(* Logix 5000 project; controller Digital_Interlock_PLC vendor 1 type 14 code 196 rev 37.11; software revision 37.00 *)

TASK MainTask (periodic, rate 10 ms, priority 5, watchdog 500 ms) : MainProgram

MODULES
   Local : vendor 1 type 14 code 196 (5069 0, rev 37.11)
      PF1 : vendor 1 type 14 code 107 (Ethernet 10.10.10.48, rev 37.1)
      ST1 : ETHERNET-MODULE (Ethernet 10.10.10.59, rev 1.1, Output RPI 10 ms)
           ST1:O.Data[0]   // To stacker heartbeat
           ST1:I.Data[1].0   // FeedInterruptStatus
      PR1 : ETHERNET-MODULE (Ethernet 10.10.10.6, rev 1.1, Output RPI 10 ms)
END_MODULES

TYPE STR_MajorFault :
STRUCT
   LEN : DINT;
   DATA : SINT[300];
END_STRUCT
END_TYPE

TYPE UDT_CommandEnum :
STRUCT
   cmd_none : DINT;
   cmd_start : DINT;
   cmd_stop : DINT;
   cmd_reset : DINT;
   cmd_interrupt : DINT;
   cmd_reconfigure : DINT;
END_STRUCT
END_TYPE

TYPE UDT_Constraints :
STRUCT
   GlobalSpeedMax : REAL;
   GlobalSpeedMin : REAL;
   KpiStabilityWindow_s : DINT;
END_STRUCT
END_TYPE

TYPE UDT_DeviceCmd :
STRUCT
   Mode : DINT;
   SpeedCmd : REAL;
   BufferTarget : DINT;
   Enable : BOOL;
END_STRUCT
END_TYPE

TYPE UDT_DeviceHealth :
STRUCT
   HeartbeatPrevious : BOOL;
   HeartbeartTimeout : BOOL;
   CommOK : BOOL;
   Enabled : BOOL;
   HeartbeatIn : BOOL;
   FaultInfo : DINT;
   EntryStatus : INT;
   FaultCode : INT;
   HBTimer : TIMER;
   Name : STRING;
   DeviceConfigured : BOOL;
END_STRUCT
END_TYPE

TYPE UDT_DeviceLink :
STRUCT
   ConnOK : BOOL;
   Simulation : BOOL;
   RoundTrip_ms : DINT;
   Handshake : UDT_Handshake;
   Cmd : UDT_DeviceCmd;
   Sts : UDT_DeviceSts;
END_STRUCT
END_TYPE

TYPE UDT_DeviceSts :
STRUCT
   PermissivesOK : BOOL;
   Running : BOOL;
   Faulted : BOOL;
   SpeedFB : REAL;
   BufferLevel : DINT;
   AlarmCode : DINT;
END_STRUCT
END_TYPE

TYPE UDT_DeviceTarget :
STRUCT
   DeviceID : DINT;
   SpeedMin : REAL;
   SpeedMax : REAL;
   BufferMin : DINT;
   BufferMax : DINT;
   Priority : DINT;
END_STRUCT
END_TYPE

TYPE UDT_EIP_DieCutter_FromStacker :   // Die cutter From Stacker
STRUCT
   blnFast : BOOL;   // Speed up die cutter (Stacker -> Press)
   blnSlow : BOOL;   // Slow down die cutter (Stacker -> Press)
   blnRegisterAdjustRq : BOOL;   // Move DC register to desired value (Stacker -> Press)
   blnRegisterStopAdjustRq : BOOL;   // Stop moving DC register (Stacker -> Press)
   blnSidewaysAdjustRq : BOOL;   // Move DC sideways to desired value (Stacker -> Press)
   blnSidewaysStopAdjustRq : BOOL;   // Stop DC sideways move (Stacker -> Press)
   blnSpeedChangeRq : BOOL;   // Change speed to desired speed (Stacker -> Press)
   blnSpeedChangeStopRq : BOOL;   // Stop speed change if active (Stacker -> Press)
   uiDesiredSpeedKpm : INT;   // 0-500 KPM (Stacker -> Press)
   fltDesiredRegisterAdjust : REAL;   // mm (Stacker -> Press)
   fltDesiredSidewaysAdjust : REAL;   // mm (Stacker -> Press)
END_STRUCT
END_TYPE

TYPE UDT_EIP_DieCutter_ToStacker :   // Die cutter to stacker
STRUCT
   blnRegistrationActive : BOOL;   // Die cutter registration motion active (Press -> Stacker)
   blnSidewaysAcitve : BOOL;   // Die cutter sideways motion active (Press -> Stacker)
   blnSpeedChangeActive : BOOL;   // Die cutter speed change active (Press -> Stacker)
   uiActualSpeedKpm : INT;   // Press current line speed (0-500 KPM) (Press -> Stacker)
   fltActualRegisterPosition : REAL;   // mm (Press -> Stacker)
   fltActualSidewaysPosition : REAL;   // mm (Press -> Stacker)
END_STRUCT
END_TYPE

TYPE UDT_EIP_FromBreaker :
STRUCT
   FeedInterrupted : BOOL;
   FeedInterrupt : BOOL;
   CurrentSpeed : DINT;
   CurrentFill : DINT;
   SampleRate : DINT;
   Deadband : DINT;
   MaxRunSpeed : DINT;
   MaxCmdSpeed : DINT;
   MinCmdSpeed : DINT;
   FeedInterruptSetting : DINT;
   TargetFill : DINT;
   CmdSpeed : DINT;
   Proportional : REAL;
   Name : STRING;
END_STRUCT
END_TYPE

TYPE UDT_EIP_FromConveyor :
STRUCT
   FeedInterrupt : BOOL;
   FeedInterrupted : BOOL;
   CurrentSpeed : DINT;
   CurrentFill : DINT;
   SampleRate : DINT;
   Deadband : DINT;
   MaxRunSpeed : DINT;
   MaxCmdSpeed : DINT;
   MinCmdSpeed : DINT;
   FeedInterruptSetting : DINT;
   TargetFill : DINT;
   CmdSpeed : DINT;
   Proportional : REAL;
   Name : STRING;
END_STRUCT
END_TYPE

TYPE UDT_EIP_FromPalletizer :
STRUCT
   FeedInterrupted : BOOL;
   FeedInterrupt : BOOL;
   CurrentSpeed : DINT;
   CurrentFill : DINT;
   SampleRate : DINT;
   Deadband : DINT;
   MaxRunSpeed : DINT;
   MaxCmdSpeed : DINT;
   MinCmdSpeed : DINT;
   FeedInterruptSetting : DINT;
   TargetFill : DINT;
   CmdSpeed : DINT;
   Proportional : REAL;
   Name : STRING;
END_STRUCT
END_TYPE

TYPE UDT_EIP_FromPrefeeder :
STRUCT
   AuxTamperAirRight : BOOL;   // (interlocks) (Pre-Feeder -> Press)
   AuxTamperAirLeft : BOOL;   // (interlocks) (Pre-Feeder -> Press)
   BackstopInhibit : BOOL;   // (Pre-Feeder -> Press)
   CallForStack : BOOL;   // Prefeeder calling for stack to be delivered (Prefeeder -> Floor Conv)
   ExtendoUpDown : BOOL;   // (interlocks) (Pre-Feeder -> Press)
   EstopFeedbackChannel1 : BOOL;   // (interlocks) (Pre-Feeder -> Press)
   EstopFeedbackChannel2 : BOOL;   // (interlocks) (Pre-Feeder -> Press)
   FeedBoardOk : BOOL;   // (interlocks) (Pre-Feeder -> Press)
   HeartbeatEcho : BOOL;
   MachineOpenCloseDisable : BOOL;   // (interlocks) (Pre-Feeder -> Press)
   OpenMachineOk : BOOL;   // (interlocks) (Pre-Feeder -> Press)
   ReadyForSetup : BOOL;   // (interlocks) (Pre-Feeder -> Press)
   ReadyToRaise : BOOL;   // (interlocks) (Pre-Feeder -> Press)
   RunEmpty : BOOL;   // (interlocks) (Pre-Feeder -> Press)
   RunForward : BOOL;   // Prefeeder telling conveyor to run forward (Prefeeder -> Floor Conv)
   RunReverse : BOOL;   // Prefeeder telling conveyor to run reverse (Prefeeder -> Floor Conv)
   TamperInterrupt : BOOL;   // (interlocks) (Pre-Feeder -> Press)
   CurrentSpeed : INT;   // Current speed of prefeeder (0-500KPM) (Pre-Feeder -> Press)
   PatternMaxSpeed : INT;   // Max speed allowed by stack pattern (0-500KPM) (Pre-Feeder -> Press)
END_STRUCT
END_TYPE

TYPE UDT_EIP_FromPress :
STRUCT
   ControlPowerInhibit : BOOL;   // Inhibit stacker from starting
   EstopOkChannel1 : BOOL;   // Press Estop is OK Ch1
   EstopOkChannel2 : BOOL;   // Press Estop is OK Ch2
   FeedEye : BOOL;   // Feed eye blocked (Press -> Stacker)
   GrinderCoverClosed : BOOL;   // OK to roll in
   LineSpeedSignal : DINT;   // Line speed of press (0-10V)
   LineEncoder : DINT;   // Enoder representing desired position of die cut cylinder rolls over every revolution (Press -> Stacker)
END_STRUCT
END_TYPE

TYPE UDT_EIP_FromStacker :
STRUCT
   ControlPower : BOOL;   // Stacker control power is on (interlocks)
   EstopOkChannel1 : BOOL;   // Stacker Estop to press ch1 (interlocks) (Stacker -> Press)
   EstopOkChannel2 : BOOL;   // Stacker Estop to press ch2 (interlocks) (Stacker -> Press)
   CompensatorControls : BOOL;   // Die Cut and Flexo Reg controls (interlocks)
   FeedInterruptStatus : BOOL;   // Interrupt request from stacker (status) (Stacker -> Press)
   FeedInterrupt : BOOL;   // Interrupt request from stacker (flow control) (Stacker -> Press)
   FeedRestart : BOOL;   // Restart feed (interlocks) (Stacker -> Press)
   HeartbeatEcho : BOOL;
   StackerRolledInChannel1 : BOOL;   // Stacker Rolled In to press Ok 2 Run Ch1 (interlocks) (Stacker -> Press)
   StackerRolledInChannel2 : BOOL;   // Stacker Rolled In to press Ok 2 Run Ch2 (interlocks) (Stacker -> Press)
   RunPermissive : BOOL;   // OK for press to run (interlocks) (Stacker -> Press)
   RolledOutStatus : BOOL;   // Die cutter rolled out (status) (Stacker -> Press)
   Spare1 : DINT;
   Spare2 : DINT;
   CurrentSpeed : INT;   // Current stacker line speed (0-500 KPM) (flow control) (Stacker -> Press)
   FillPercentage : INT;   // Percentage of Accumulation Consumed (for calculating Upstream Machine Speed) (flow control) (Stacker -> Press)
   PatternMaxSpeed : INT;   // Maximum speed allowed by stacker pattern (0-500 KPM) (flow control) (Stacker -> Press)
   Heartbeat : UINT;   // Heartbeat Reflection from Stacker (interlocks) (Stacker -> Press)
   DieCutter : UDT_EIP_DieCutter_FromStacker;
   PrintStation : UDT_EIP_PrintStation_FromStacker[7];
END_STRUCT
END_TYPE

TYPE UDT_EIP_FromStrapper :
STRUCT
   FeedInterrupt : BOOL;
   FeedInterrupted : BOOL;
   CurrentSpeed : DINT;
   CurrentFill : DINT;
   SampleRate : DINT;
   Deadband : DINT;
   MaxRunSpeed : DINT;
   MaxCmdSpeed : DINT;
   MinCmdSpeed : DINT;
   FeedInterruptSetting : DINT;
   TargetFill : DINT;
   CmdSpeed : DINT;
   Proportional : REAL;
   Name : STRING;
END_STRUCT
END_TYPE

TYPE UDT_EIP_FromTwinBoxSlitter :
STRUCT
   FeedInterrupt : BOOL;
   FeedInterrupted : BOOL;
   CurrentSpeed : DINT;
   CurrentFill : DINT;
   SampleRate : DINT;
   Deadband : DINT;
   MaxRunSpeed : DINT;
   MaxCmdSpeed : DINT;
   MinCmdSpeed : DINT;
   FeedInterruptSetting : DINT;
   TargetFill : DINT;
   CmdSpeed : DINT;
   Proportional : REAL;
   Name : STRING;
END_STRUCT
END_TYPE

TYPE UDT_EIP_PrintStation_FromStacker :   // print station from stacker
STRUCT
   blnRegisterAdjustRq : BOOL;   // (Stacker -> Press)
   blnSidewaysAdjustRq : BOOL;   // (Stacker -> Press)
   blnRegisterStopAdjustRq : BOOL;   // (Stacker -> Press)
   blnSidewaysStopAdjustRq : BOOL;   // (Stacker -> Press)
   fltDesiredRegisterAdjust : REAL;   // mm (Stacker -> Press)
   fltDesiredSidewaysAdjust : REAL;   // mm (Stacker -> Press)
END_STRUCT
END_TYPE

TYPE UDT_EIP_PrintStation_ToStacker :   // print station to stacker
STRUCT
   blnRegistrationActive : BOOL;   // (Press -> Stacker)
   blnSideWaysActive : BOOL;   // (Press -> Stacker)
   fltActualRegisterPosition : REAL;   // mm (Press -> Stacker)
   fltActualSidewaysPosition : REAL;   // mm (Press -> Stacker)
END_STRUCT
END_TYPE

TYPE UDT_EIP_ToBreaker :
STRUCT
   FeedInterrupted : BOOL;
   FeedInterrupt : BOOL;
   CurrentSpeed : DINT;
   CurrentFill : DINT;
   SampleRate : DINT;
   Deadband : DINT;
   MaxRunSpeed : DINT;
   MaxCmdSpeed : DINT;
   MinCmdSpeed : DINT;
   FeedInterruptSetting : DINT;
   TargetFill : DINT;
   CmdSpeed : DINT;
   Proportional : REAL;
   Name : STRING;
END_STRUCT
END_TYPE

TYPE UDT_EIP_ToConveyor :
STRUCT
   FeedInterrupt : BOOL;
   FeedInterrupted : BOOL;
   CurrentSpeed : DINT;
   CurrentFill : DINT;
   SampleRate : DINT;
   Deadband : DINT;
   MaxRunSpeed : DINT;
   MaxCmdSpeed : DINT;
   MinCmdSpeed : DINT;
   FeedInterruptSetting : DINT;
   TargetFill : DINT;
   CmdSpeed : DINT;
   Proportional : REAL;
   Name : STRING;
END_STRUCT
END_TYPE

TYPE UDT_EIP_ToPalletizer :
STRUCT
   FeedInterrupted : BOOL;
   FeedInterrupt : BOOL;
   CurrentSpeed : DINT;
   CurrentFill : DINT;
   SampleRate : DINT;
   Deadband : DINT;
   MaxRunSpeed : DINT;
   MaxCmdSpeed : DINT;
   MinCmdSpeed : DINT;
   FeedInterruptSetting : DINT;
   TargetFill : DINT;
   CmdSpeed : DINT;
   Proportional : REAL;
   Name : STRING;
END_STRUCT
END_TYPE

TYPE UDT_EIP_ToPrefeeder :
STRUCT
   ClosedLocked : BOOL;   // (interlocks) (Press -> Pre-Feeder)
   ConvRunning : BOOL;   // (Floor Conv -> Prefeeder)
   ExtendoFollowBackstopUp : BOOL;   // (interlocks) (Press -> Pre-Feeder)
   ExtendoFollowBackstopDown : BOOL;   // (interlocks) (Press -> Pre-Feeder)
   LastStack : BOOL;   // Last stack running in (Floor Conv -> Prefeeder)
   LoadHopper : BOOL;   // (interlocks) (Press -> Pre-Feeder)
   MachineInFeedMode : BOOL;   // (interlocks) (Press -> Pre-Feeder)
   MachineRunning : BOOL;   // (interlocks) (Press -> Pre-Feeder)
   RequestsOpen : BOOL;   // (interlocks) (Press -> Pre-Feeder)
   StackReadyInFeed : BOOL;   // Stack is present at the end of the floor conveyor (Floor Conv -> Prefeeder)
   ShuttleCarAtPrefeeder : BOOL;   // (Floor Conv -> Prefeeder)
   Heartbeat : DINT;
   CommandedSpeed : INT;   // Commanded speed from the Press/LIC (0-500KPM) (flow control) (Press -> Pre-Feeder)
   BoardCaliper : REAL;   // Thickness of board (mm) (interlocks) (Press -> Pre-Feeder)
   FeedHopperHeight : REAL;   // (mm) (interlocks) (Press -> Pre-Feeder)
   HopperHeightSetpoint : REAL;   // (mm) (interlocks) (Press -> Pre-Feeder)
   HopperHeightMin : REAL;   // (mm) (interlocks) (Press -> Pre-Feeder)
   LinearSpeedSetpoint : REAL;   // Setting based on recipe (mm/s) (interlocks) (Press -> Pre-Feeder)
   LinearSpeedActual : REAL;   // Actual speed (mm/s) (interlocks) (Press -> Pre-Feeder)
END_STRUCT
END_TYPE

TYPE UDT_EIP_ToPress :
STRUCT
   AuxTamperAirRight : BOOL;   // (Pre-Feeder -> Press)
   AuxTamperAirLeft : BOOL;   // (Pre-Feeder -> Press)
   CallForStack : BOOL;   // Prefeeder -> Floor Conv
   FeedBoardOk : BOOL;   // (Pre-Feeder -> Press)
   MachineOpenCloseDisable : BOOL;   // (Pre-Feeder -> Press)
   OpenMachineOk : BOOL;   // (Pre-Feeder -> Press)
   ReadyForSetup : BOOL;   // (Pre-Feeder -> Press)
   ReadyToRaise : BOOL;   // (Pre-Feeder -> Press)
   RunEmpty : BOOL;
   RunForward : BOOL;   // (Pre-Feeder -> Press)
   RunReverse : BOOL;   // (Pre-Feeder -> Press)
   TamperInterrupt : BOOL;   // (Pre-Feeder -> Press)
   Empty : BOOL;   // (Pre-Feeder -> Press)
   BackstopInhibit : BOOL;   // (Prefeeder -> Press)
   Placeholder : BOOL;
   FeedInterrupt : BOOL;   // Interrupt request from stacker (flow control)
   FeedRestart : BOOL;   // Restart feed (interlocks)
   EstopFeedbackChannel1 : BOOL;   // (Prefeeder -> Press)
   EstopFeedbackChannel2 : BOOL;   // (Prefeeder -> Press)
   EstopOkChannel1 : BOOL;   // Stacker Estop to press ch1 (interlocks)
   EstopOkChannel2 : BOOL;   // Stacker Estop to press ch2 (interlocks)
   ExtendoUpDown : BOOL;   // (interlocks) (Pre-Feeder -> Press)
   StackerRolledInChannel1 : BOOL;   // Stacker Rolled In to press Ok 2 Run Ch1 (interlocks)
   StackerRolledInChannel2 : BOOL;   // Stacker Rolled In to press Ok 2 Run Ch2 (interlocks)
   ControlPower : BOOL;   // Stacker control power is on (interlocks)
   CompensatorControls : BOOL;   // Die Cut and Flexo Reg controls (interlocks)
   RunPermissive : BOOL;   // OK for press to run (interlocks)
   RolledOutStatus : BOOL;   // Die cutter rolled out (status)
   FeedInterruptStatus : BOOL;   // Interrupt request from stacker (status)
   Spare : BOOL;
   Heartbeat_Echo_Prefeeder : UINT;   // Heartbeat Reflection from Prefeeder (interlocks) (Prefeeder -> Press)
   Heartbeat_Echo_Stacker : UINT;   // Heartbeat Reflection from Stacker (interlocks) (Stacker -> Press)
   CurrentSpeed : UINT;   // Current stacker line speed (0-500 KPM) (flow control) (Pre-Feeder -> Press)
   PatternMaxSpeed : UINT;   // Maximum speed allowed by stacker pattern (0-500 KPM) (flow control) (Pre-Feeder -> Press)
   FillPercentage : UINT;   // Percentage of Accumulation Consumed (for calculating Upstream Machine Speed) (flow control)
   Spare1 : DINT;
   Spare2 : DINT;
   DieCutter : UDT_EIP_DieCutter_ToStacker;
   PrintStation : UDT_EIP_PrintStation_FromStacker[7];
END_STRUCT
END_TYPE

TYPE UDT_EIP_ToStacker :
STRUCT
   ControlPowerInhibit : BOOL;   // ADDED FOR EIP COMMS Inhibit stacker from starting
   DownstreamReady : BOOL;   // (LIC -> Stacker)
   EstopOkChannel1 : BOOL;   // Press Estop is OK Ch1 (interlocks) (Press -> Stacker)
   EstopOkChannel2 : BOOL;   // Press Estop is OK Ch2 (interlocks) (Press -> Stacker)
   FeedEye : BOOL;   // ADDED FOR EIP COMMS Feed eye blocked
   GrinderCoverClosed : BOOL;   // ADDED FOR EIP COMMS OK to roll in
   RollInPermissive : BOOL;   // Permission for stacker roll-in (Press -> Stacker)
   RunPermissive : BOOL;   // Rum permissive from press (interlocks) (Press -> Stacker)
   SheetCountPulseStatus : BOOL;   // Sheet count pulse (interlocks) (Press -> Stacker)
   VOSReset : BOOL;   // Reset VOS faults (if applicable) (interlocks) (Press -> Stacker)
   VOSStart : BOOL;   // Start VOS (if applicable) (interlocks) (Press -> Stacker)
   CommsStatus : DINT;   // (Interlock -> Stacker)
   Spare1 : DINT;
   Spare2 : DINT;
   LineEncoder : DINT;   // ADDED FOR EIP COMMS Enoder representing desired position of die cut cylinder rolls over every revolution
   LineSpeedSignal : DINT;   // ADDED FOR EIP COMMS Line speed of press (0-10V)
   CommandedSpeed : INT;   // Commanded press speed (0-500 KPM) (Press -> Stacker)
   PressCurrentSpeed : INT;   // Actual press speed (0-500 KPM) (Press -> Stacker)
   Heartbeat : UINT;   // Incrementing heartbeat for comm health (Press -> Stacker)
   DieCutter : UDT_EIP_DieCutter_ToStacker;
   PrintStation : UDT_EIP_PrintStation_ToStacker[7];
END_STRUCT
END_TYPE

TYPE UDT_EIP_ToStrapper :
STRUCT
   FeedInterrupt : BOOL;
   FeedInterrupted : BOOL;
   CurrentSpeed : DINT;
   CurrentFill : DINT;
   SampleRate : DINT;
   Deadband : DINT;
   MaxRunSpeed : DINT;
   MaxCmdSpeed : DINT;
   MinCmdSpeed : DINT;
   FeedInterruptSetting : DINT;
   TargetFill : DINT;
   CmdSpeed : DINT;
   Proportional : REAL;
   Name : STRING;
END_STRUCT
END_TYPE

TYPE UDT_EIP_ToTwinBoxSlitter :
STRUCT
   FeedInterrupt : BOOL;
   FeedInterrupted : BOOL;
   CurrentSpeed : DINT;
   CurrentFill : DINT;
   SampleRate : DINT;
   Deadband : DINT;
   MaxRunSpeed : DINT;
   MaxCmdSpeed : DINT;
   MinCmdSpeed : DINT;
   FeedInterruptSetting : DINT;
   TargetFill : DINT;
   CmdSpeed : DINT;
   Proportional : REAL;
   Name : STRING;
END_STRUCT
END_TYPE

TYPE UDT_FaultRecord :
STRUCT
   TimeLow : DINT;
   TimeHigh : DINT;
   Type : INT;
   Code : INT;
   Info : DINT[11];
END_STRUCT
END_TYPE

TYPE UDT_FromLIC :   // Data that is exchanged with LIC Client
STRUCT
   EnableLineOptimization : BOOL;
   Deadband : DINT;
   FeedInterruptSetting : DINT;
   MaxCommandSpeed : DINT;
   MinCommandSpeed : DINT;
   Proportional : DINT;
   SampleRate : DINT;
   TargetFillPercentage : DINT;
   MachineList : STRING;
   ToBR1 : UDT_EIP_ToBreaker;
   ToBR2 : UDT_EIP_ToBreaker;
   ToCN1 : UDT_EIP_ToConveyor;
   ToCN2 : UDT_EIP_ToConveyor;
   ToPL1 : UDT_EIP_ToPalletizer;
   ToPL2 : UDT_EIP_ToPalletizer;
   ToFE1 : UDT_EIP_ToPrefeeder;
   ToFE2 : UDT_EIP_ToPrefeeder;
   ToPR1 : UDT_EIP_ToPress;
   ToPR2 : UDT_EIP_ToPress;
   ToST1 : UDT_EIP_ToStacker;
   ToST2 : UDT_EIP_ToStacker;
   ToTB1 : UDT_EIP_ToTwinBoxSlitter;
   ToTB2 : UDT_EIP_ToTwinBoxSlitter;
   ToSR1 : UDT_EIP_ToStrapper;
   ToSR2 : UDT_EIP_ToStrapper;
END_STRUCT
END_TYPE

TYPE UDT_GenericStacker :
STRUCT
   cmd : DINT;
   status : DINT;
END_STRUCT
END_TYPE

TYPE UDT_Handshake :   // Device handshake and telemetry
STRUCT
   Req : BOOL;
   Ack : BOOL;
   Busy : BOOL;
   Done : BOOL;
   Fault : BOOL;
   TxnID : DINT;
   TxnIDEcho : DINT;
   Timeout_ms : DINT;
   Timer_ms : DINT;
END_STRUCT
END_TYPE

TYPE UDT_MachineType :
STRUCT
   ModuleExists : BOOL;   // (Handled by SetModuleInhibitMode) A bool that represents unihibited (0,False) or inhibited (1,True)
   FeedInterrupt : BOOL;   // (Output to each PLC) Boolean for activating feed interrupt
   FeedInterrupted : BOOL;   // Flag to verify feed interrupt execution
   ProportialGain : REAL;   // Proportial multiple to adjust aggressiveness of changes to speed commands, limited to [0.5 - 1.2]
   MachineType : STRING;   // (From HMI) List of configured machines, with format "FE1,PR1,SR1,ST1,PL1"
   CurrentSpeed : DINT;   // (From each PLC) Each machine will have a current speed value, obtained over EIP
   MinSpeed : DINT;   // (From each PLC) Minimum speed of the machine
   CommandSpeed : DINT;   // (Output of Line Flow Opt) Commanded speed adjustment from speed algorithm, occurs every *evaluation interval*
   IPSubnet : DINT;   // (**CHECK** if HMI will provide) The subnet that maps to the type of machine
   FeedInterruptSetting : DINT;   // (Input from HMI) Value from 0 to 100% , above which the press feed interrupt is triggered
   ReferenceSpeed : DINT;   // (Obtained from reference list, derived from machine list) Speed reference of downstream machine
   CurrFillPercentage : DINT;   // (From each PLC) Fill percentage of current machine
   TargFillPercentage : DINT;   // (From HMI per machine) The target fill percentage that is used to calculate commanded speeds
   Deadband : DINT;   // Value that represents the amount of percentage points from target fill percentage that the current fill percentage must be before calculating command speed
   MaxCmdSpeed : DINT;   // (From HMI) Value in KPM representing the upper limit of the commanded speed to be output to the upstream machine
   MinCmdSpeed : DINT;   // (From HMI) Value in KPM representing the lower limit of the commanded speed to be output to the upstream machine
END_STRUCT
END_TYPE

TYPE UDT_Optimize_Command :
STRUCT
   Enable : BOOL;
   Request : BOOL;
   Cancel : BOOL;
   Reset : BOOL;
END_STRUCT
END_TYPE

TYPE UDT_Optimize_Config :
STRUCT
   RecipeID : DINT;
   Mode : DINT;
   Targets : UDT_DeviceTarget[15];
   Constraints : UDT_Constraints;
END_STRUCT
END_TYPE

TYPE UDT_Optimize_Status :
STRUCT
   Active : BOOL;
   Busy : BOOL;
   Complete : BOOL;
   Fault : BOOL;
   Step : DINT;
   Substep : DINT;
   TimeInState_ms : DINT;
   LastErrorCode : DINT;
   LastErrorText : DINT;
   TxnID : DINT;
END_STRUCT
END_TYPE

TYPE UDT_StateContext :
STRUCT
   AbortReq : BOOL;
   Alarm : BOOL;
   Busy : BOOL;
   Complete : BOOL;
   InitDone : BOOL;
   StateChanged : BOOL;
   StartRisingEdge : BOOL;
   StopRisingEdge : BOOL;
   ResetRisingEdge : BOOL;
   PreviousStart : BOOL;
   PreviousStop : BOOL;
   PreviousReset : BOOL;
   InterruptRisingEdge : BOOL;
   PreviousInterrupt : BOOL;
   PreviousDone : BOOL;
   DoneRisingEdge : BOOL;
   Previous : DINT;
   Current : DINT;
   EntryStamp : DINT;   // ms since power-up
   TimeInState_ms : DINT;
   Command : DINT;   // from HMI/mailbox
   CommandID : DINT;   // monotonic; prevents replays
   Fault : DINT;   // 0 = none; otherwise code
   Next : DINT;
END_STRUCT
END_TYPE

TYPE UDT_States :
STRUCT
   IDLE : DINT;
   INITIALIZE : DINT;
   RUNNING : DINT;
   STOPPING : DINT;
   FAULT : DINT;
   ERROR : DINT;
   COMPLETE : DINT;
   INTERRUPT : DINT;
   HOLD : DINT;
   STARTING : DINT;
END_STRUCT
END_TYPE

TYPE UDT_ToLIC :
STRUCT
   FeedInterrupt : BOOL;   // Feed interrupt executed
   FeedInterrupted : BOOL;   // Interrupt completed
   CommsHealthy : BOOL;   // All machines are communicating
   MachinesConnected : BOOL[32];   // Boolean array that contains machine connection status
   FromBR1 : UDT_EIP_FromBreaker;
   FromBR2 : UDT_EIP_FromBreaker;
   FromCN1 : UDT_EIP_FromConveyor;
   FromCN2 : UDT_EIP_FromConveyor;
   FromPL1 : UDT_EIP_FromPalletizer;
   FromPL2 : UDT_EIP_FromPalletizer;
   FromFE1 : UDT_EIP_FromPrefeeder;
   FromFE2 : UDT_EIP_FromPrefeeder;
   FromPR1 : UDT_EIP_FromPress;
   FromPR2 : UDT_EIP_FromPress;
   FromST1 : UDT_EIP_FromStacker;
   FromST2 : UDT_EIP_FromStacker;
   FromTB1 : UDT_EIP_FromTwinBoxSlitter;
   FromTB2 : UDT_EIP_FromTwinBoxSlitter;
   FromSR1 : UDT_EIP_FromStrapper;
   FromSR2 : UDT_EIP_FromStrapper;
END_STRUCT
END_TYPE

ADD_ON_INSTRUCTION AOI_EIP_DEVICE   (* revision 1.0 *)
VAR_INPUT
   Inp_Inhibit : BOOL;
   Inp_PermissivesOK : BOOL;
END_VAR
VAR_IN_OUT
   Inp_Cmd : UDT_DeviceCmd; {required}
END_VAR
VAR_INPUT
   Inp_ReqSetpoint : BOOL;
   Inp_TxnID : DINT;
   Inp_Timeout_ms : DINT;
END_VAR
VAR_IN_OUT
   Line : UDT_DeviceLink; {required}
END_VAR
VAR_OUTPUT
   Out_Succeeded : BOOL; {access Read Only}
   Out_Faulted : BOOL; {access Read Only}
   Out_Verified : BOOL; {access Read Only}
END_VAR

ROUTINE Logic   (* structured text *)
   
END_ROUTINE
END_ADD_ON_INSTRUCTION

ADD_ON_INSTRUCTION AOI_LineFlowOptimization   (* revision 1.0 *)
// Line Speed Adjustment
VAR_INPUT
   CurrSpeed : DINT; {required}   // Current speed of the target machine (KPM)
END_VAR
VAR_OUTPUT
   CmdSpeed : DINT; {required}   // The command speed output by the speed alrgothim, written to target machine (KPM)
END_VAR
VAR_INPUT
   RefSpeed : DINT; {required}   // Reference speed of the downstream machine (KPM)
   CurrFillPer : DINT; {required}   // Current Fill Percentage (%) of consumed buffer capacity
   TargFillPer : DINT; {required}   // Target Fill Percentage, the desired fill percentage to achieve by adjusting speeds (%)
   MaxSpeed : DINT; {required}   // Maximum speed of job (KPM)
   MinSpeed : DINT; {required}   // Minimum speed of target machine (KPM)
END_VAR
VAR_OUTPUT
   FeedInterrupt : BOOL; {required}   // Value set to TRUE, when the Reference Fill % is equal to or greater than the Feed Interrupt Setting LIC Client user input).
END_VAR
VAR_INPUT
   FeedInterruptSetting : DINT; {required}   // Value set by LIC Client user interface
   SpeedEvalRate : DINT; {required}   // Rate of speed calculations
END_VAR
VAR
   FillPerTimer : TIMER;
   ProportionalGain : DINT;   // Proportial multiple to adjust aggressiveness of changes to speed commands, limited to [0.5 - 1.2]
   DeadBand : DINT;   // Value that represents the amount of percentage points from target fill percentage that the current fill percentage must be before calculating command speed
   LowDBand : DINT;
   HighDBand : DINT;
END_VAR

ROUTINE Logic   (* ladder *)
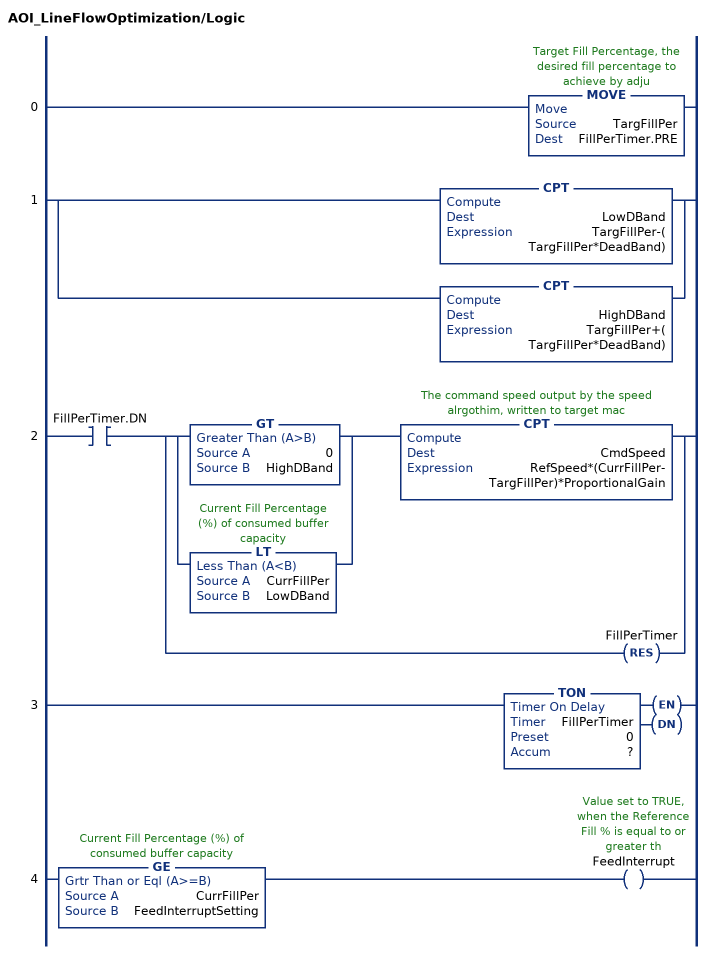
   0: MOVE(TargFillPer,FillPerTimer.PRE);
   1: [CPT(LowDBand,TargFillPer-(TargFillPer*DeadBand)) ,CPT(HighDBand,TargFillPer+(TargFillPer*DeadBand)) ];
   2: XIC(FillPerTimer.DN)[[GT(0,HighDBand) ,LT(CurrFillPer,LowDBand) ] CPT(CmdSpeed,RefSpeed*(CurrFillPer-TargFillPer)*ProportionalGain) ,RES(FillPerTimer) ];
   3: TON(FillPerTimer,?,?);
   4: GE(CurrFillPer,FeedInterruptSetting)OTE(FeedInterrupt);
END_ROUTINE
END_ADD_ON_INSTRUCTION

ADD_ON_INSTRUCTION AOI_ModuleInhibitManager   (* revision 1.0 *)
// Accepts a list of allowed module names (array of strings) and a count. Modules in the list are uninhibited and modules not included are inhibited. Intended for a project with up to MAX_MODULES generic Ethernet modules (default 16). Designed non-blocking and deterministic: call once per request or on a periodic task.
VAR_IN_OUT
   Inp_ConfiguredList : STRING; {required}
END_VAR
VAR_INPUT
   Inp_ConfiguredCount : DINT;   // Number of configured machines in list
END_VAR
VAR_OUTPUT
   Out_Done : BOOL; {access Read Only}
   Out_Error : BOOL; {access Read Only}
   Out_ErrorCode : DINT; {access Read Only}
   Out_UpdatedCount : DINT; {access Read Only}   // number of modules changed (for diagnostics)
END_VAR
VAR_INPUT
   Inp_Execute : BOOL;
   Inp_MaxModules : DINT;
END_VAR
VAR
   Configured16 : STRING[16]; {access None}
   Configured15 : STRING[15]; {access None}
   Configured14 : STRING[14]; {access None}
   Configured13 : STRING[13]; {access None}
   Configured12 : STRING[12]; {access None}
   Configured11 : STRING[11]; {access None}
   Configured10 : STRING[10]; {access None}
   Configured9 : STRING[9]; {access None}
   Configured8 : STRING[8]; {access None}
   Configured7 : STRING[7]; {access None}
   Configured6 : STRING[6]; {access None}
   Configured5 : STRING[5]; {access None}
   Configured4 : STRING[4]; {access None}
   out : STRING; {access None}
   i : DINT; {access None}
   changes : DINT; {access None}
   stagedInhibit : BOOL[32]; {access None}
   cmpAllowedName : STRING; {access None}
   cmpModuleName : STRING; {access None}
   prevExecute : BOOL; {access None}
   found : BOOL; {access None}
   j : DINT; {access None}
   maxMachAllowed : DINT := 16; {access None}
END_VAR

ROUTINE Logic   (* structured text *)
// Accepts a list of allowed module names (array of strings) and a count. Modules in the list are uninhibited and modules not included are inhibited. Intended for a project with up to MAX_MODULES generic Ethernet modules (default 16). Designed non-blocking and deterministic: call once per request or on a periodic task.
   (* Initialize outputs each scan;
   Done will be latched until Execute clears (design choice) *)
   Out_Done := 0;
   Out_Error := 0;
   Out_ErrorCode := 0;
   Out_UpdatedCount := 0;
   (*Validate inputs*)
   if (Inp_ConfiguredCount < 0) OR (Inp_ConfiguredCount > maxMachAllowed) then
   	Out_Error := 1;
   	Out_ErrorCode := -1; (* Invalid machine count*)
   end_if;
   
   if (Inp_MaxModules < 1) OR (Inp_MaxModules > maxMachAllowed) then
   	Out_Error := 1;
   	Out_ErrorCode := 2; (* Invalid MaxModules*)
   end_if;
   
   (* Rising-edge detect (if you prefer Execute to be pulse). If you want Execute held to reflect active,
   remove the prevExecute check and run update whenever Execute is TRUE. *)
   if Inp_Execute AND NOT prevExecute then
   	(* Build stagedInhibit[]: default to TRUE (inhibit) then clear for matches *)
   	for i := 1 to Inp_MaxModules do
   		stagedInhibit[i] := 1; (* assume inhibited unless found in allowed list *)
   	end_for;
   
      (* For each configured module, search the AllowedList *)
   	changes := 0;
   	for i:= 1 to Inp_MaxModules do
   		(* Safety: empty module names are considered not allowed / inhibited *)
   		if Inp_ConfiguredList.LEN = 0 then
   			stagedInhibit[i] := 1;
   		end_if;
   		found := 0;
   		for j := 1 to Inp_ConfiguredCount do
   			if Inp_ConfiguredList.LEN = 0 then
   			end_if;
   		end_for;
   	end_for;
   end_if;
   
   
   
   
   
END_ROUTINE
END_ADD_ON_INSTRUCTION

ADD_ON_INSTRUCTION AOI_OPT_STATE   (* revision 1.0 *)

ROUTINE Logic   (* structured text *)
   
END_ROUTINE
END_ADD_ON_INSTRUCTION

ADD_ON_INSTRUCTION AOI_Optimize   (* revision 1.0 *)
VAR_INPUT
   Inp_CurrentFill : DINT; {required}   // Current Fill Percentage (%) of consumed buffer capacity
   Inp_CurrentSpeed : DINT; {required}   // Current speed of the target machine (KPM)
   Inp_FeedInterruptSetting : DINT; {required}   // Value set by LIC Client user interface
   Inp_MaxSpeed : DINT; {required}   // Maximum speed of job (KPM)
   Inp_MinSpeed : DINT; {required}   // Minimum speed of target machine (KPM)
   Inp_ReferenceSpeed : DINT; {required}   // Reference speed of the downstream machine (KPM)
   Inp_SamplingRate : DINT; {required}   // Rate of speed calculations
   Inp_TargetFill : DINT; {required}   // Target Fill Percentage, the desired fill percentage to achieve by adjusting speeds (%)
END_VAR
VAR_OUTPUT
   Out_CommandSpeed : DINT; {required}   // The command speed output by the speed alrgothim, written to target machine (KPM)
   Out_FeedInterrupt : BOOL; {required}   // Value set to TRUE, when the Reference Fill % is equal to or greater than the Feed Interrupt Setting LIC Client user input).
END_VAR
VAR
   FillTimer : TIMER := (PRE := 500);
   Inp_Deadband : DINT;   // Value that represents the amount of percentage points from target fill percentage that the current fill percentage must be before calculating command speed
   Inp_ProportionalGain : DINT;   // Proportial multiple to adjust aggressiveness of changes to speed commands, limited to [0.5 - 1.2]
   LowerDeadband : DINT;
   UpperDeadband : DINT;
END_VAR

ROUTINE Logic   (* structured text *)
   //Configure timer
   FillTimer.PRE := 500;
   
   //Calculate deadband limits
   LowerDeadband := Inp_TargetFill - (Inp_TargetFill * Inp_Deadband);
   UpperDeadband := Inp_TargetFill + (Inp_TargetFill * Inp_Deadband);
   
   //After each cycle of the Fill Timer, check if the current fill percentage is outside the
   //deadband bounds, compute command speed if it is.
   if (FillTimer.DN) then
   	if (Inp_CurrentFill > UpperDeadband) OR (Inp_CurrentFill < LowerDeadband) then
   		//The command speed output by the speed alrgothim, written to target machine (KPM)
   		Out_CommandSpeed := Inp_ReferenceSpeed * (Inp_CurrentFill - Inp_TargetFill) * Inp_ProportionalGain;
   	end_if;
   
   	// Explicit reset for timer
   	FillTimer.EN := 0;
   	FillTimer.EN := 1;
   end_if;
   
   //Enable Timer
   FillTimer.EN := 1;
   
   //If current fill exceeds feed interrupt setting, initiate Feed interrupt
   if (Inp_CurrentFill >= Inp_FeedInterruptSetting) then
   	Out_FeedInterrupt := 1;
   end_if;
   
END_ROUTINE
END_ADD_ON_INSTRUCTION

ADD_ON_INSTRUCTION AOI_ResetMachineArray   (* revision 1.0 *)
VAR_IN_OUT
   Inp_Machine : UDT_MachineType; {required}
END_VAR

ROUTINE Logic   (* structured text *)
   Inp_Machine.CommandSpeed 			:= 0;
   Inp_Machine.CurrentSpeed 			:= 0;
   Inp_Machine.CurrFillPercentage 		:= 0;
   Inp_Machine.Deadband 				:= 0;
   Inp_Machine.FeedInterrupt 			:= 0;
   Inp_Machine.FeedInterrupted			:= 0;
   Inp_Machine.FeedInterruptSetting 	:= 0;
   Inp_Machine.IPSubnet 				:= 0;
   Inp_Machine.MachineType 			:= '';
   Inp_Machine.MaxCmdSpeed 			:= 0;
   Inp_Machine.MinCmdSpeed 			:= 0;
   Inp_Machine.MinCmdSpeed 			:= 0;
   Inp_Machine.MinSpeed 				:= 0;
   Inp_Machine.ModuleExists 			:= 0;
   Inp_Machine.ProportialGain 			:= 0;
   Inp_Machine.ReferenceSpeed 			:= 0;
   Inp_Machine.TargFillPercentage 		:= 0;
END_ROUTINE
END_ADD_ON_INSTRUCTION
